   "Carrier_46_SpareInput(4_6)" AT %I2666.6 : Bool;   // SPARE INPUT
   "Carrier_46_SpareInput(4_7)" AT %I2666.7 : Bool;   // SPARE INPUT
   "Carrier_46_PB1_ProdHoldLH" AT %I2667.0 : Bool;   // PB 1 PRODUCTION HOLD LH
   "Carrier_46_PB2_ResetLH" AT %I2667.1 : Bool;   // PB 2 RESET LH
   "Carrier_46_PB3_ProdHoldRH" AT %I2667.2 : Bool;   // PB 3 PRODUCTION HOLD RH
   "Carrier_46_PB4_ResetRH" AT %I2667.3 : Bool;   // PB 4 RESET RH
   "Carrier_46_SpareInput(4_14)" AT %I2667.4 : Bool;   // SPARE INPUT
   "Carrier_46_SpareInput(4_15)" AT %I2667.5 : Bool;   // SPARE INPUT
   "Carrier_46_SpareInput(4_16)" AT %I2667.6 : Bool;   // SPARE INPUT
   "Carrier_46_SpareInput(4_17)" AT %I2667.7 : Bool;   // SPARE INPUT
   "Carrier_46_Slot5_Output" AT %IW2668 : Word;   // SLOT 5 OUTPUT WORD
   "Carrier_46_IRD400_HMI_24VDC_ENABLE" AT %I2668.0 : Bool;   // IRD 400 PANEL HMI 24V DC POWER
   "Carrier_46_FaultLight_LH" AT %I2668.1 : Bool;   // FAULT LIGHT LH
   "Carrier_46_RunLight_LH" AT %I2668.2 : Bool;   // RUN LIGHT LH
   "Carrier_46_FaultLight_RH" AT %I2668.3 : Bool;   // FAULT LIGHT RH
   "Carrier_46_RunLight_RH" AT %I2668.4 : Bool;   // RUN LIGHT RH
   "Carrier_46_SpareOutput(5_5)" AT %I2668.5 : Bool;   // SPARE OUTPUT
   "Carrier_46_SpareOutput(5_6)" AT %I2668.6 : Bool;   // SPARE OUTPUT
   "Carrier_46_SpareOutput(5_7)" AT %I2668.7 : Bool;   // SPARE OUTPUT
   "Carrier_46_ActualSpeed" AT %IW2670 : Word;   // ACTUAL SPEED
   "Carrier_46_CarrierDriveAlarm" AT %IW2672 : Word;   // CARRIER DRIVE ALARM
   "Carrier_46_CarrierDriveWarning" AT %IW2674 : Word;   // CARRIER DRIVE WARNING
   "Carrier_47_Status" AT %IW2700 : Word;   // CARRIER STATUS WORD
   "Carrier_47_Status.0" AT %I2700.0 : Bool;   // HEARTBEAT
   "Carrier_47_Status.1" AT %I2700.1 : Bool;   // MANUAL
   "Carrier_47_Status.2" AT %I2700.2 : Bool;   // IN_AUTO
   "Carrier_47_Status.3" AT %I2700.3 : Bool;   // POSITIONING_COMPLETE
   "Carrier_47_Status.4" AT %I2700.4 : Bool;   // PRODUCTION HOLD
   "Carrier_47_Status.5" AT %I2700.5 : Bool;   // CARRIER MOVING FORWARD
   "Carrier_47_Status.6" AT %I2700.6 : Bool;   // CARRIER MOVING REVERSE
   "Carrier_47_Status.7" AT %I2700.7 : Bool;   // CARRIER FAULT
   "Carrier_47_Status.8" AT %I2701.0 : Bool;   // CRASH DETECT TRIPPED
   "Carrier_47_Status.9" AT %I2701.1 : Bool;
   "Carrier_47_Status.10" AT %I2701.2 : Bool;
   "Carrier_47_Status.11" AT %I2701.3 : Bool;
   "Carrier_47_Status.12" AT %I2701.4 : Bool;
   "Carrier_47_Status.13" AT %I2701.5 : Bool;
   "Carrier_47_Status.14" AT %I2701.6 : Bool;
   "Carrier_47_Status.15" AT %I2701.7 : Bool;
   "Carrier_47_SDCFaultCode" AT %IW2702 : Word;   // SDC FAULT CODE
   "Carrier_47_CarrierPosition" AT %ID2704 : DWord;   // CARRIER POSITION
   "Carrier_47_CarrierNumber" AT %IW2708 : Word;   // CARRIER NUMBER
   "Carrier_47_G120DControlWord" AT %IW2710 : Word;   // G120D_STW1_CONTROL
   "Carrier_47_G120DControlWord.0" AT %I2710.0 : Bool;   // Bit_00_ON
   "Carrier_47_G120DControlWord.1" AT %I2710.1 : Bool;   // Bit_01_AUS2_INH
   "Carrier_47_G120DControlWord.2" AT %I2710.2 : Bool;   // Bit_02_AUS3_STOP
   "Carrier_47_G120DControlWord.3" AT %I2710.3 : Bool;   // Bit_03_EN
   "Carrier_47_G120DControlWord.4" AT %I2710.4 : Bool;   // Bit_04_EN_RAMP
   "Carrier_47_G120DControlWord.5" AT %I2710.5 : Bool;   // Bit_05_START_RAMP
   "Carrier_47_G120DControlWord.6" AT %I2710.6 : Bool;   // Bit_06_SETPOINT
   "Carrier_47_G120DControlWord.7" AT %I2710.7 : Bool;   // Bit_07_RESET
   "Carrier_47_G120DControlWord.8" AT %I2711.0 : Bool;   // Bit_08_JOG_R
   "Carrier_47_G120DControlWord.9" AT %I2711.1 : Bool;   // Bit_09_JOG_L
   "Carrier_47_G120DControlWord.10" AT %I2711.2 : Bool;   // Bit_10_CONTR_PLC
   "Carrier_47_G120DControlWord.11" AT %I2711.3 : Bool;   // Bit_11_REVERSE
   "Carrier_47_G120DControlWord.12" AT %I2711.4 : Bool;   // Bit_12_BRAKE_RELEASE
   "Carrier_47_G120DControlWord.13" AT %I2711.5 : Bool;   // Bit_13_DDS
   "Carrier_47_G120DControlWord.14" AT %I2711.6 : Bool;   // Bit_14_DO0
   "Carrier_47_G120DControlWord.15" AT %I2711.7 : Bool;   // Bit_15_DO1
   "Carrier_47_G120DStatusWord" AT %IW2712 : Word;   // G120D_ZSW1_STATUS
   "Carrier_47_G120DStatusWord.0" AT %I2712.0 : Bool;   // Bit_00_READY_RUN
   "Carrier_47_G120DStatusWord.1" AT %I2712.1 : Bool;   // Bit_01_READY_ON
   "Carrier_47_G120DStatusWord.2" AT %I2712.2 : Bool;   // Bit_02_ENABLE
   "Carrier_47_G120DStatusWord.3" AT %I2712.3 : Bool;   // Bit_03_FAULT
   "Carrier_47_G120DStatusWord.4" AT %I2712.4 : Bool;   // Bit_04_OFF2
   "Carrier_47_G120DStatusWord.5" AT %I2712.5 : Bool;   // Bit_05_OFF3
   "Carrier_47_G120DStatusWord.6" AT %I2712.6 : Bool;   // Bit_06_LOCK_OUT
   "Carrier_47_G120DStatusWord.7" AT %I2712.7 : Bool;   // Bit_07_WARN
   "Carrier_47_G120DStatusWord.8" AT %I2713.0 : Bool;   // Bit_08_NO_DEVIATION
   "Carrier_47_G120DStatusWord.9" AT %I2713.1 : Bool;   // Bit_09_CONTR_PLC
   "Carrier_47_G120DStatusWord.10" AT %I2713.2 : Bool;   // Bit_10_F_MAX
   "Carrier_47_G120DStatusWord.11" AT %I2713.3 : Bool;   // Bit_11_LIMIT_REACHED
   "Carrier_47_G120DStatusWord.12" AT %I2713.4 : Bool;   // Bit_12_BRAKE_OPEN
   "Carrier_47_G120DStatusWord.13" AT %I2713.5 : Bool;   // Bit_13_NO_OVERTEMP
   "Carrier_47_G120DStatusWord.14" AT %I2713.6 : Bool;   // Bit_14_CW_CCW
   "Carrier_47_G120DStatusWord.15" AT %I2713.7 : Bool;   // Bit_15_OVERL
   "Carrier_47_Slot2_Input" AT %IW2714 : Word;   // SLOT 2 INPUT WORD
   "Carrier_47_CrashDetectSW" AT %I2714.0 : Bool;   // CRASH DETECT SW
   "Carrier_47_SpareSafetyInput(2_1)" AT %I2714.1 : Bool;   // SPARE SAFETY INPUT
   "Carrier_47_SpareSafetyInput(2_2)" AT %I2714.2 : Bool;   // SPARE SAFETY INPUT
   "Carrier_47_SpareSafetyInput(2_3)" AT %I2714.3 : Bool;   // SPARE SAFETY INPUT
   "Carrier_47_SpareSafetyInput(2_4)" AT %I2714.4 : Bool;   // SPARE SAFETY INPUT
   "Carrier_47_SpareSafetyInput(2_5)" AT %I2714.5 : Bool;   // SPARE SAFETY INPUT
   "Carrier_47_SpareSafetyInput(2_6)" AT %I2714.6 : Bool;   // SPARE SAFETY INPUT
   "Carrier_47_SpareSafetyInput(2_7)" AT %I2714.7 : Bool;   // SPARE SAFETY INPUT
   "Carrier_47_Slot3_SafetyOutput" AT %IW2715 : Word;   // SLOT 3 SAFETY OUTPUT WORD
   "Carrier_47_Crash_Detect_OK" AT %I2715.0 : Bool;   // CARRIER CRASH DETECT
   "Carrier_47_SpareSafetyOutput(3_1)" AT %I2715.1 : Bool;   // SPARE SAFETY OUTPUT
   "Carrier_47_SpareSafetyOutput(3_2)" AT %I2715.2 : Bool;   // SPARE SAFETY OUTPUT
   "Carrier_47_SpareSafetyOutput(3_3)" AT %I2715.3 : Bool;   // SPARE SAFETY OUTPUT
   "Carrier_47_SpareSafetyOutput(3_4)" AT %I2715.4 : Bool;   // SPARE SAFETY OUTPUT
   "Carrier_47_SpareSafetyOutput(3_5)" AT %I2715.5 : Bool;   // SPARE SAFETY OUTPUT
   "Carrier_47_SpareSafetyOutput(3_6)" AT %I2715.6 : Bool;   // SPARE SAFETY OUTPUT
   "Carrier_47_SpareSafetyOutput(3_7)" AT %I2715.7 : Bool;   // SPARE SAFETY OUTPUT
   "Carrier_47_Slot4_Input" AT %IW2716 : Word;   // SLOT 4 INPUT WORD
   "Carrier_47_480VPowerOn_MDCB1" AT %I2716.0 : Bool;   // 480 VAC POWER ON MDCB 1
   "Carrier_47_SpareInput(4_1)" AT %I2716.1 : Bool;   // SPARE INPUT
   "Carrier_47_SpareInput(4_2)" AT %I2716.2 : Bool;   // SPARE INPUT
   "Carrier_47_SitopSelectStatus" AT %I2716.3 : Bool;   // SITOP SELECT STATUS
   "Carrier_47_DCsupplyOnPSCB2" AT %I2716.4 : Bool;   // DC SUPPLY ON PSCB 2
   "Carrier_47_SpareInput(4_5)" AT %I2716.5 : Bool;   // SPARE INPUT
   "Carrier_47_SpareInput(4_6)" AT %I2716.6 : Bool;   // SPARE INPUT
   "Carrier_47_SpareInput(4_7)" AT %I2716.7 : Bool;   // SPARE INPUT
   "Carrier_47_PB1_ProdHoldLH" AT %I2717.0 : Bool;   // PB 1 PRODUCTION HOLD LH
   "Carrier_47_PB2_ResetLH" AT %I2717.1 : Bool;   // PB 2 RESET LH
   "Carrier_47_PB3_ProdHoldRH" AT %I2717.2 : Bool;   // PB 3 PRODUCTION HOLD RH
   "Carrier_47_PB4_ResetRH" AT %I2717.3 : Bool;   // PB 4 RESET RH
   "Carrier_47_SpareInput(4_14)" AT %I2717.4 : Bool;   // SPARE INPUT
   "Carrier_47_SpareInput(4_15)" AT %I2717.5 : Bool;   // SPARE INPUT
   "Carrier_47_SpareInput(4_16)" AT %I2717.6 : Bool;   // SPARE INPUT
   "Carrier_47_SpareInput(4_17)" AT %I2717.7 : Bool;   // SPARE INPUT
   "Carrier_47_Slot5_Output" AT %IW2718 : Word;   // SLOT 5 OUTPUT WORD
   "Carrier_47_IRD400_HMI_24VDC_ENABLE" AT %I2718.0 : Bool;   // IRD 400 PANEL HMI 24V DC POWER
   "Carrier_47_FaultLight_LH" AT %I2718.1 : Bool;   // FAULT LIGHT LH
   "Carrier_47_RunLight_LH" AT %I2718.2 : Bool;   // RUN LIGHT LH
   "Carrier_47_FaultLight_RH" AT %I2718.3 : Bool;   // FAULT LIGHT RH
   "Carrier_47_RunLight_RH" AT %I2718.4 : Bool;   // RUN LIGHT RH
   "Carrier_47_SpareOutput(5_5)" AT %I2718.5 : Bool;   // SPARE OUTPUT
   "Carrier_47_SpareOutput(5_6)" AT %I2718.6 : Bool;   // SPARE OUTPUT
   "Carrier_47_SpareOutput(5_7)" AT %I2718.7 : Bool;   // SPARE OUTPUT
   "Carrier_47_ActualSpeed" AT %IW2720 : Word;   // ACTUAL SPEED
   "Carrier_47_CarrierDriveAlarm" AT %IW2722 : Word;   // CARRIER DRIVE ALARM
   "Carrier_47_CarrierDriveWarning" AT %IW2724 : Word;   // CARRIER DRIVE WARNING
   "Carrier_48_Status" AT %IW2750 : Word;   // CARRIER STATUS WORD
   "Carrier_48_Status.0" AT %I2750.0 : Bool;   // HEARTBEAT
   "Carrier_48_Status.1" AT %I2750.1 : Bool;   // MANUAL
   "Carrier_48_Status.2" AT %I2750.2 : Bool;   // IN_AUTO
   "Carrier_48_Status.3" AT %I2750.3 : Bool;   // POSITIONING_COMPLETE
   "Carrier_48_Status.4" AT %I2750.4 : Bool;   // PRODUCTION HOLD
   "Carrier_48_Status.5" AT %I2750.5 : Bool;   // CARRIER MOVING FORWARD
   "Carrier_48_Status.6" AT %I2750.6 : Bool;   // CARRIER MOVING REVERSE
   "Carrier_48_Status.7" AT %I2750.7 : Bool;   // CARRIER FAULT
   "Carrier_48_Status.8" AT %I2751.0 : Bool;   // CRASH DETECT TRIPPED
   "Carrier_48_Status.9" AT %I2751.1 : Bool;
   "Carrier_48_Status.10" AT %I2751.2 : Bool;
   "Carrier_48_Status.11" AT %I2751.3 : Bool;
   "Carrier_48_Status.12" AT %I2751.4 : Bool;
   "Carrier_48_Status.13" AT %I2751.5 : Bool;
   "Carrier_48_Status.14" AT %I2751.6 : Bool;
   "Carrier_48_Status.15" AT %I2751.7 : Bool;
   "Carrier_48_SDCFaultCode" AT %IW2752 : Word;   // SDC FAULT CODE
   "Carrier_48_CarrierPosition" AT %ID2754 : DWord;   // CARRIER POSITION
   "Carrier_48_CarrierNumber" AT %IW2758 : Word;   // CARRIER NUMBER
   "Carrier_48_G120DControlWord" AT %IW2760 : Word;   // G120D_STW1_CONTROL
   "Carrier_48_G120DControlWord.0" AT %I2760.0 : Bool;   // Bit_00_ON
   "Carrier_48_G120DControlWord.1" AT %I2760.1 : Bool;   // Bit_01_AUS2_INH
   "Carrier_48_G120DControlWord.2" AT %I2760.2 : Bool;   // Bit_02_AUS3_STOP
   "Carrier_48_G120DControlWord.3" AT %I2760.3 : Bool;   // Bit_03_EN
   "Carrier_48_G120DControlWord.4" AT %I2760.4 : Bool;   // Bit_04_EN_RAMP
   "Carrier_48_G120DControlWord.5" AT %I2760.5 : Bool;   // Bit_05_START_RAMP
   "Carrier_48_G120DControlWord.6" AT %I2760.6 : Bool;   // Bit_06_SETPOINT
   "Carrier_48_G120DControlWord.7" AT %I2760.7 : Bool;   // Bit_07_RESET
   "Carrier_48_G120DControlWord.8" AT %I2761.0 : Bool;   // Bit_08_JOG_R
   "Carrier_48_G120DControlWord.9" AT %I2761.1 : Bool;   // Bit_09_JOG_L
   "Carrier_48_G120DControlWord.10" AT %I2761.2 : Bool;   // Bit_10_CONTR_PLC
   "Carrier_48_G120DControlWord.11" AT %I2761.3 : Bool;   // Bit_11_REVERSE
   "Carrier_48_G120DControlWord.12" AT %I2761.4 : Bool;   // Bit_12_BRAKE_RELEASE
   "Carrier_48_G120DControlWord.13" AT %I2761.5 : Bool;   // Bit_13_DDS
   "Carrier_48_G120DControlWord.14" AT %I2761.6 : Bool;   // Bit_14_DO0
   "Carrier_48_G120DControlWord.15" AT %I2761.7 : Bool;   // Bit_15_DO1
   "Carrier_48_G120DStatusWord" AT %IW2762 : Word;   // G120D_ZSW1_STATUS
   "Carrier_48_G120DStatusWord.0" AT %I2762.0 : Bool;   // Bit_00_READY_RUN
   "Carrier_48_G120DStatusWord.1" AT %I2762.1 : Bool;   // Bit_01_READY_ON
   "Carrier_48_G120DStatusWord.2" AT %I2762.2 : Bool;   // Bit_02_ENABLE
   "Carrier_48_G120DStatusWord.3" AT %I2762.3 : Bool;   // Bit_03_FAULT
   "Carrier_48_G120DStatusWord.4" AT %I2762.4 : Bool;   // Bit_04_OFF2
   "Carrier_48_G120DStatusWord.5" AT %I2762.5 : Bool;   // Bit_05_OFF3
   "Carrier_48_G120DStatusWord.6" AT %I2762.6 : Bool;   // Bit_06_LOCK_OUT
   "Carrier_48_G120DStatusWord.7" AT %I2762.7 : Bool;   // Bit_07_WARN
   "Carrier_48_G120DStatusWord.8" AT %I2763.0 : Bool;   // Bit_08_NO_DEVIATION
   "Carrier_48_G120DStatusWord.9" AT %I2763.1 : Bool;   // Bit_09_CONTR_PLC
   "Carrier_48_G120DStatusWord.10" AT %I2763.2 : Bool;   // Bit_10_F_MAX
   "Carrier_48_G120DStatusWord.11" AT %I2763.3 : Bool;   // Bit_11_LIMIT_REACHED
   "Carrier_48_G120DStatusWord.12" AT %I2763.4 : Bool;   // Bit_12_BRAKE_OPEN
   "Carrier_48_G120DStatusWord.13" AT %I2763.5 : Bool;   // Bit_13_NO_OVERTEMP
   "Carrier_48_G120DStatusWord.14" AT %I2763.6 : Bool;   // Bit_14_CW_CCW
   "Carrier_48_G120DStatusWord.15" AT %I2763.7 : Bool;   // Bit_15_OVERL
   "Carrier_48_Slot2_Input" AT %IW2764 : Word;   // SLOT 2 INPUT WORD
   "Carrier_48_CrashDetectSW" AT %I2764.0 : Bool;   // CRASH DETECT SW
   "Carrier_48_SpareSafetyInput(2_1)" AT %I2764.1 : Bool;   // SPARE SAFETY INPUT
   "Carrier_48_SpareSafetyInput(2_2)" AT %I2764.2 : Bool;   // SPARE SAFETY INPUT
   "Carrier_48_SpareSafetyInput(2_3)" AT %I2764.3 : Bool;   // SPARE SAFETY INPUT
   "Carrier_48_SpareSafetyInput(2_4)" AT %I2764.4 : Bool;   // SPARE SAFETY INPUT
   "Carrier_48_SpareSafetyInput(2_5)" AT %I2764.5 : Bool;   // SPARE SAFETY INPUT
   "Carrier_48_SpareSafetyInput(2_6)" AT %I2764.6 : Bool;   // SPARE SAFETY INPUT
   "Carrier_48_SpareSafetyInput(2_7)" AT %I2764.7 : Bool;   // SPARE SAFETY INPUT
   "Carrier_48_Slot3_SafetyOutput" AT %IW2765 : Word;   // SLOT 3 SAFETY OUTPUT WORD
   "Carrier_48_Crash_Detect_OK" AT %I2765.0 : Bool;   // CARRIER CRASH DETECT
   "Carrier_48_SpareSafetyOutput(3_1)" AT %I2765.1 : Bool;   // SPARE SAFETY OUTPUT
   "Carrier_48_SpareSafetyOutput(3_2)" AT %I2765.2 : Bool;   // SPARE SAFETY OUTPUT
   "Carrier_48_SpareSafetyOutput(3_3)" AT %I2765.3 : Bool;   // SPARE SAFETY OUTPUT
   "Carrier_48_SpareSafetyOutput(3_4)" AT %I2765.4 : Bool;   // SPARE SAFETY OUTPUT
   "Carrier_48_SpareSafetyOutput(3_5)" AT %I2765.5 : Bool;   // SPARE SAFETY OUTPUT
   "Carrier_48_SpareSafetyOutput(3_6)" AT %I2765.6 : Bool;   // SPARE SAFETY OUTPUT
   "Carrier_48_SpareSafetyOutput(3_7)" AT %I2765.7 : Bool;   // SPARE SAFETY OUTPUT
   "Carrier_48_Slot4_Input" AT %IW2766 : Word;   // SLOT 4 INPUT WORD
   "Carrier_48_480VPowerOn_MDCB1" AT %I2766.0 : Bool;   // 480 VAC POWER ON MDCB 1
   "Carrier_48_SpareInput(4_1)" AT %I2766.1 : Bool;   // SPARE INPUT
   "Carrier_48_SpareInput(4_2)" AT %I2766.2 : Bool;   // SPARE INPUT
   "Carrier_48_SitopSelectStatus" AT %I2766.3 : Bool;   // SITOP SELECT STATUS
   "Carrier_48_DCsupplyOnPSCB2" AT %I2766.4 : Bool;   // DC SUPPLY ON PSCB 2
   "Carrier_48_SpareInput(4_5)" AT %I2766.5 : Bool;   // SPARE INPUT
   "Carrier_48_SpareInput(4_6)" AT %I2766.6 : Bool;   // SPARE INPUT
   "Carrier_48_SpareInput(4_7)" AT %I2766.7 : Bool;   // SPARE INPUT
   "Carrier_48_PB1_ProdHoldLH" AT %I2767.0 : Bool;   // PB 1 PRODUCTION HOLD LH
   "Carrier_48_PB2_ResetLH" AT %I2767.1 : Bool;   // PB 2 RESET LH
   "Carrier_48_PB3_ProdHoldRH" AT %I2767.2 : Bool;   // PB 3 PRODUCTION HOLD RH
   "Carrier_48_PB4_ResetRH" AT %I2767.3 : Bool;   // PB 4 RESET RH
   "Carrier_48_SpareInput(4_14)" AT %I2767.4 : Bool;   // SPARE INPUT
   "Carrier_48_SpareInput(4_15)" AT %I2767.5 : Bool;   // SPARE INPUT
   "Carrier_48_SpareInput(4_16)" AT %I2767.6 : Bool;   // SPARE INPUT
   "Carrier_48_SpareInput(4_17)" AT %I2767.7 : Bool;   // SPARE INPUT
   "Carrier_48_Slot5_Output" AT %IW2768 : Word;   // SLOT 5 OUTPUT WORD
   "Carrier_48_IRD400_HMI_24VDC_ENABLE" AT %I2768.0 : Bool;   // IRD 400 PANEL HMI 24V DC POWER
   "Carrier_48_FaultLight_LH" AT %I2768.1 : Bool;   // FAULT LIGHT LH
   "Carrier_48_RunLight_LH" AT %I2768.2 : Bool;   // RUN LIGHT LH
   "Carrier_48_FaultLight_RH" AT %I2768.3 : Bool;   // FAULT LIGHT RH
   "Carrier_48_RunLight_RH" AT %I2768.4 : Bool;   // RUN LIGHT RH
   "Carrier_48_SpareOutput(5_5)" AT %I2768.5 : Bool;   // SPARE OUTPUT
   "Carrier_48_SpareOutput(5_6)" AT %I2768.6 : Bool;   // SPARE OUTPUT
   "Carrier_48_SpareOutput(5_7)" AT %I2768.7 : Bool;   // SPARE OUTPUT
   "Carrier_48_ActualSpeed" AT %IW2770 : Word;   // ACTUAL SPEED
   "Carrier_48_CarrierDriveAlarm" AT %IW2772 : Word;   // CARRIER DRIVE ALARM
   "Carrier_48_CarrierDriveWarning" AT %IW2774 : Word;   // CARRIER DRIVE WARNING
   "Carrier_49_Status" AT %IW2800 : Word;   // CARRIER STATUS WORD
   "Carrier_49_Status.0" AT %I2800.0 : Bool;   // HEARTBEAT
   "Carrier_49_Status.1" AT %I2800.1 : Bool;   // MANUAL
   "Carrier_49_Status.2" AT %I2800.2 : Bool;   // IN_AUTO
   "Carrier_49_Status.3" AT %I2800.3 : Bool;   // POSITIONING_COMPLETE
   "Carrier_49_Status.4" AT %I2800.4 : Bool;   // PRODUCTION HOLD
   "Carrier_49_Status.5" AT %I2800.5 : Bool;   // CARRIER MOVING FORWARD
   "Carrier_49_Status.6" AT %I2800.6 : Bool;   // CARRIER MOVING REVERSE
   "Carrier_49_Status.7" AT %I2800.7 : Bool;   // CARRIER FAULT
   "Carrier_49_Status.8" AT %I2801.0 : Bool;   // CRASH DETECT TRIPPED
   "Carrier_49_Status.9" AT %I2801.1 : Bool;
   "Carrier_49_Status.10" AT %I2801.2 : Bool;
   "Carrier_49_Status.11" AT %I2801.3 : Bool;
   "Carrier_49_Status.12" AT %I2801.4 : Bool;
   "Carrier_49_Status.13" AT %I2801.5 : Bool;
   "Carrier_49_Status.14" AT %I2801.6 : Bool;
   "Carrier_49_Status.15" AT %I2801.7 : Bool;
   "Carrier_49_SDCFaultCode" AT %IW2802 : Word;   // SDC FAULT CODE
   "Carrier_49_CarrierPosition" AT %ID2804 : DWord;   // CARRIER POSITION
   "Carrier_49_CarrierNumber" AT %IW2808 : Word;   // CARRIER NUMBER
   "Carrier_49_G120DControlWord" AT %IW2810 : Word;   // G120D_STW1_CONTROL
   "Carrier_49_G120DControlWord.0" AT %I2810.0 : Bool;   // Bit_00_ON
   "Carrier_49_G120DControlWord.1" AT %I2810.1 : Bool;   // Bit_01_AUS2_INH
   "Carrier_49_G120DControlWord.2" AT %I2810.2 : Bool;   // Bit_02_AUS3_STOP
   "Carrier_49_G120DControlWord.3" AT %I2810.3 : Bool;   // Bit_03_EN
   "Carrier_49_G120DControlWord.4" AT %I2810.4 : Bool;   // Bit_04_EN_RAMP
   "Carrier_49_G120DControlWord.5" AT %I2810.5 : Bool;   // Bit_05_START_RAMP
   "Carrier_49_G120DControlWord.6" AT %I2810.6 : Bool;   // Bit_06_SETPOINT
   "Carrier_49_G120DControlWord.7" AT %I2810.7 : Bool;   // Bit_07_RESET
   "Carrier_49_G120DControlWord.8" AT %I2811.0 : Bool;   // Bit_08_JOG_R
   "Carrier_49_G120DControlWord.9" AT %I2811.1 : Bool;   // Bit_09_JOG_L
   "Carrier_49_G120DControlWord.10" AT %I2811.2 : Bool;   // Bit_10_CONTR_PLC
   "Carrier_49_G120DControlWord.11" AT %I2811.3 : Bool;   // Bit_11_REVERSE
   "Carrier_49_G120DControlWord.12" AT %I2811.4 : Bool;   // Bit_12_BRAKE_RELEASE
   "Carrier_49_G120DControlWord.13" AT %I2811.5 : Bool;   // Bit_13_DDS
   "Carrier_49_G120DControlWord.14" AT %I2811.6 : Bool;   // Bit_14_DO0
   "Carrier_49_G120DControlWord.15" AT %I2811.7 : Bool;   // Bit_15_DO1
   "Carrier_49_G120DStatusWord" AT %IW2812 : Word;   // G120D_ZSW1_STATUS
   "Carrier_49_G120DStatusWord.0" AT %I2812.0 : Bool;   // Bit_00_READY_RUN
   "Carrier_49_G120DStatusWord.1" AT %I2812.1 : Bool;   // Bit_01_READY_ON
   "Carrier_49_G120DStatusWord.2" AT %I2812.2 : Bool;   // Bit_02_ENABLE
   "Carrier_49_G120DStatusWord.3" AT %I2812.3 : Bool;   // Bit_03_FAULT
   "Carrier_49_G120DStatusWord.4" AT %I2812.4 : Bool;   // Bit_04_OFF2
   "Carrier_49_G120DStatusWord.5" AT %I2812.5 : Bool;   // Bit_05_OFF3
   "Carrier_49_G120DStatusWord.6" AT %I2812.6 : Bool;   // Bit_06_LOCK_OUT
   "Carrier_49_G120DStatusWord.7" AT %I2812.7 : Bool;   // Bit_07_WARN
   "Carrier_49_G120DStatusWord.8" AT %I2813.0 : Bool;   // Bit_08_NO_DEVIATION
   "Carrier_49_G120DStatusWord.9" AT %I2813.1 : Bool;   // Bit_09_CONTR_PLC
   "Carrier_49_G120DStatusWord.10" AT %I2813.2 : Bool;   // Bit_10_F_MAX
   "Carrier_49_G120DStatusWord.11" AT %I2813.3 : Bool;   // Bit_11_LIMIT_REACHED
   "Carrier_49_G120DStatusWord.12" AT %I2813.4 : Bool;   // Bit_12_BRAKE_OPEN
   "Carrier_49_G120DStatusWord.13" AT %I2813.5 : Bool;   // Bit_13_NO_OVERTEMP
   "Carrier_49_G120DStatusWord.14" AT %I2813.6 : Bool;   // Bit_14_CW_CCW
   "Carrier_49_G120DStatusWord.15" AT %I2813.7 : Bool;   // Bit_15_OVERL
   "Carrier_49_Slot2_Input" AT %IW2814 : Word;   // SLOT 2 INPUT WORD
   "Carrier_49_CrashDetectSW" AT %I2814.0 : Bool;   // CRASH DETECT SW
   "Carrier_49_SpareSafetyInput(2_1)" AT %I2814.1 : Bool;   // SPARE SAFETY INPUT
   "Carrier_49_SpareSafetyInput(2_2)" AT %I2814.2 : Bool;   // SPARE SAFETY INPUT
   "Carrier_49_SpareSafetyInput(2_3)" AT %I2814.3 : Bool;   // SPARE SAFETY INPUT
   "Carrier_49_SpareSafetyInput(2_4)" AT %I2814.4 : Bool;   // SPARE SAFETY INPUT
   "Carrier_49_SpareSafetyInput(2_5)" AT %I2814.5 : Bool;   // SPARE SAFETY INPUT
   "Carrier_49_SpareSafetyInput(2_6)" AT %I2814.6 : Bool;   // SPARE SAFETY INPUT
   "Carrier_49_SpareSafetyInput(2_7)" AT %I2814.7 : Bool;   // SPARE SAFETY INPUT
   "Carrier_49_Slot3_SafetyOutput" AT %IW2815 : Word;   // SLOT 3 SAFETY OUTPUT WORD
   "Carrier_49_Crash_Detect_OK" AT %I2815.0 : Bool;   // CARRIER CRASH DETECT
   "Carrier_49_SpareSafetyOutput(3_1)" AT %I2815.1 : Bool;   // SPARE SAFETY OUTPUT
   "Carrier_49_SpareSafetyOutput(3_2)" AT %I2815.2 : Bool;   // SPARE SAFETY OUTPUT
   "Carrier_49_SpareSafetyOutput(3_3)" AT %I2815.3 : Bool;   // SPARE SAFETY OUTPUT
   "Carrier_49_SpareSafetyOutput(3_4)" AT %I2815.4 : Bool;   // SPARE SAFETY OUTPUT
   "Carrier_49_SpareSafetyOutput(3_5)" AT %I2815.5 : Bool;   // SPARE SAFETY OUTPUT
   "Carrier_49_SpareSafetyOutput(3_6)" AT %I2815.6 : Bool;   // SPARE SAFETY OUTPUT
   "Carrier_49_SpareSafetyOutput(3_7)" AT %I2815.7 : Bool;   // SPARE SAFETY OUTPUT
   "Carrier_49_Slot4_Input" AT %IW2816 : Word;   // SLOT 4 INPUT WORD
   "Carrier_49_480VPowerOn_MDCB1" AT %I2816.0 : Bool;   // 480 VAC POWER ON MDCB 1
   "Carrier_49_SpareInput(4_1)" AT %I2816.1 : Bool;   // SPARE INPUT
   "Carrier_49_SpareInput(4_2)" AT %I2816.2 : Bool;   // SPARE INPUT
   "Carrier_49_SitopSelectStatus" AT %I2816.3 : Bool;   // SITOP SELECT STATUS
   "Carrier_49_DCsupplyOnPSCB2" AT %I2816.4 : Bool;   // DC SUPPLY ON PSCB 2
   "Carrier_49_SpareInput(4_5)" AT %I2816.5 : Bool;   // SPARE INPUT
   "Carrier_49_SpareInput(4_6)" AT %I2816.6 : Bool;   // SPARE INPUT
   "Carrier_49_SpareInput(4_7)" AT %I2816.7 : Bool;   // SPARE INPUT
   "Carrier_49_PB1_ProdHoldLH" AT %I2817.0 : Bool;   // PB 1 PRODUCTION HOLD LH
   "Carrier_49_PB2_ResetLH" AT %I2817.1 : Bool;   // PB 2 RESET LH
   "Carrier_49_PB3_ProdHoldRH" AT %I2817.2 : Bool;   // PB 3 PRODUCTION HOLD RH
   "Carrier_49_PB4_ResetRH" AT %I2817.3 : Bool;   // PB 4 RESET RH
   "Carrier_49_SpareInput(4_14)" AT %I2817.4 : Bool;   // SPARE INPUT
   "Carrier_49_SpareInput(4_15)" AT %I2817.5 : Bool;   // SPARE INPUT
   "Carrier_49_SpareInput(4_16)" AT %I2817.6 : Bool;   // SPARE INPUT
   "Carrier_49_SpareInput(4_17)" AT %I2817.7 : Bool;   // SPARE INPUT
   "Carrier_49_Slot5_Output" AT %IW2818 : Word;   // SLOT 5 OUTPUT WORD
   "Carrier_49_IRD400_HMI_24VDC_ENABLE" AT %I2818.0 : Bool;   // IRD 400 PANEL HMI 24V DC POWER
   "Carrier_49_FaultLight_LH" AT %I2818.1 : Bool;   // FAULT LIGHT LH
   "Carrier_49_RunLight_LH" AT %I2818.2 : Bool;   // RUN LIGHT LH
   "Carrier_49_FaultLight_RH" AT %I2818.3 : Bool;   // FAULT LIGHT RH
   "Carrier_49_RunLight_RH" AT %I2818.4 : Bool;   // RUN LIGHT RH
   "Carrier_49_SpareOutput(5_5)" AT %I2818.5 : Bool;   // SPARE OUTPUT
   "Carrier_49_SpareOutput(5_6)" AT %I2818.6 : Bool;   // SPARE OUTPUT
   "Carrier_49_SpareOutput(5_7)" AT %I2818.7 : Bool;   // SPARE OUTPUT
   "Carrier_49_ActualSpeed" AT %IW2820 : Word;   // ACTUAL SPEED
   "Carrier_49_CarrierDriveAlarm" AT %IW2822 : Word;   // CARRIER DRIVE ALARM
   "Carrier_49_CarrierDriveWarning" AT %IW2824 : Word;   // CARRIER DRIVE WARNING
   "Carrier_50_Status" AT %IW2850 : Word;   // CARRIER STATUS WORD
   "Carrier_50_Status.0" AT %I2850.0 : Bool;   // HEARTBEAT
   "Carrier_50_Status.1" AT %I2850.1 : Bool;   // MANUAL
   "Carrier_50_Status.2" AT %I2850.2 : Bool;   // IN_AUTO
   "Carrier_50_Status.3" AT %I2850.3 : Bool;   // POSITIONING_COMPLETE
   "Carrier_50_Status.4" AT %I2850.4 : Bool;   // PRODUCTION HOLD
   "Carrier_50_Status.5" AT %I2850.5 : Bool;   // CARRIER MOVING FORWARD
   "Carrier_50_Status.6" AT %I2850.6 : Bool;   // CARRIER MOVING REVERSE
   "Carrier_50_Status.7" AT %I2850.7 : Bool;   // CARRIER FAULT
   "Carrier_50_Status.8" AT %I2851.0 : Bool;   // CRASH DETECT TRIPPED
   "Carrier_50_Status.9" AT %I2851.1 : Bool;
   "Carrier_50_Status.10" AT %I2851.2 : Bool;
   "Carrier_50_Status.11" AT %I2851.3 : Bool;
   "Carrier_50_Status.12" AT %I2851.4 : Bool;
   "Carrier_50_Status.13" AT %I2851.5 : Bool;
   "Carrier_50_Status.14" AT %I2851.6 : Bool;
   "Carrier_50_Status.15" AT %I2851.7 : Bool;
   "Carrier_50_SDCFaultCode" AT %IW2852 : Word;   // SDC FAULT CODE
   "Carrier_50_CarrierPosition" AT %ID2854 : DWord;   // CARRIER POSITION
   "Carrier_50_CarrierNumber" AT %IW2858 : Word;   // CARRIER NUMBER
   "Carrier_50_G120DControlWord" AT %IW2860 : Word;   // G120D_STW1_CONTROL
   "Carrier_50_G120DControlWord.0" AT %I2860.0 : Bool;   // Bit_00_ON
   "Carrier_50_G120DControlWord.1" AT %I2860.1 : Bool;   // Bit_01_AUS2_INH
   "Carrier_50_G120DControlWord.2" AT %I2860.2 : Bool;   // Bit_02_AUS3_STOP
   "Carrier_50_G120DControlWord.3" AT %I2860.3 : Bool;   // Bit_03_EN
   "Carrier_50_G120DControlWord.4" AT %I2860.4 : Bool;   // Bit_04_EN_RAMP
   "Carrier_50_G120DControlWord.5" AT %I2860.5 : Bool;   // Bit_05_START_RAMP
   "Carrier_50_G120DControlWord.6" AT %I2860.6 : Bool;   // Bit_06_SETPOINT
   "Carrier_50_G120DControlWord.7" AT %I2860.7 : Bool;   // Bit_07_RESET
   "Carrier_50_G120DControlWord.8" AT %I2861.0 : Bool;   // Bit_08_JOG_R
   "Carrier_50_G120DControlWord.9" AT %I2861.1 : Bool;   // Bit_09_JOG_L
   "Carrier_50_G120DControlWord.10" AT %I2861.2 : Bool;   // Bit_10_CONTR_PLC
   "Carrier_50_G120DControlWord.11" AT %I2861.3 : Bool;   // Bit_11_REVERSE
   "Carrier_50_G120DControlWord.12" AT %I2861.4 : Bool;   // Bit_12_BRAKE_RELEASE
   "Carrier_50_G120DControlWord.13" AT %I2861.5 : Bool;   // Bit_13_DDS
   "Carrier_50_G120DControlWord.14" AT %I2861.6 : Bool;   // Bit_14_DO0
   "Carrier_50_G120DControlWord.15" AT %I2861.7 : Bool;   // Bit_15_DO1
   "Carrier_50_G120DStatusWord" AT %IW2862 : Word;   // G120D_ZSW1_STATUS
   "Carrier_50_G120DStatusWord.0" AT %I2862.0 : Bool;   // Bit_00_READY_RUN
   "Carrier_50_G120DStatusWord.1" AT %I2862.1 : Bool;   // Bit_01_READY_ON
   "Carrier_50_G120DStatusWord.2" AT %I2862.2 : Bool;   // Bit_02_ENABLE
   "Carrier_50_G120DStatusWord.3" AT %I2862.3 : Bool;   // Bit_03_FAULT
   "Carrier_50_G120DStatusWord.4" AT %I2862.4 : Bool;   // Bit_04_OFF2
   "Carrier_50_G120DStatusWord.5" AT %I2862.5 : Bool;   // Bit_05_OFF3
   "Carrier_50_G120DStatusWord.6" AT %I2862.6 : Bool;   // Bit_06_LOCK_OUT
   "Carrier_50_G120DStatusWord.7" AT %I2862.7 : Bool;   // Bit_07_WARN
   "Carrier_50_G120DStatusWord.8" AT %I2863.0 : Bool;   // Bit_08_NO_DEVIATION
   "Carrier_50_G120DStatusWord.9" AT %I2863.1 : Bool;   // Bit_09_CONTR_PLC
   "Carrier_50_G120DStatusWord.10" AT %I2863.2 : Bool;   // Bit_10_F_MAX
   "Carrier_50_G120DStatusWord.11" AT %I2863.3 : Bool;   // Bit_11_LIMIT_REACHED
   "Carrier_50_G120DStatusWord.12" AT %I2863.4 : Bool;   // Bit_12_BRAKE_OPEN
   "Carrier_50_G120DStatusWord.13" AT %I2863.5 : Bool;   // Bit_13_NO_OVERTEMP
   "Carrier_50_G120DStatusWord.14" AT %I2863.6 : Bool;   // Bit_14_CW_CCW
   "Carrier_50_G120DStatusWord.15" AT %I2863.7 : Bool;   // Bit_15_OVERL
   "Carrier_50_Slot2_Input" AT %IW2864 : Word;   // SLOT 2 INPUT WORD
   "Carrier_50_CrashDetectSW" AT %I2864.0 : Bool;   // CRASH DETECT SW
   "Carrier_50_SpareSafetyInput(2_1)" AT %I2864.1 : Bool;   // SPARE SAFETY INPUT
   "Carrier_50_SpareSafetyInput(2_2)" AT %I2864.2 : Bool;   // SPARE SAFETY INPUT
   "Carrier_50_SpareSafetyInput(2_3)" AT %I2864.3 : Bool;   // SPARE SAFETY INPUT
   "Carrier_50_SpareSafetyInput(2_4)" AT %I2864.4 : Bool;   // SPARE SAFETY INPUT
   "Carrier_50_SpareSafetyInput(2_5)" AT %I2864.5 : Bool;   // SPARE SAFETY INPUT
   "Carrier_50_SpareSafetyInput(2_6)" AT %I2864.6 : Bool;   // SPARE SAFETY INPUT
   "Carrier_50_SpareSafetyInput(2_7)" AT %I2864.7 : Bool;   // SPARE SAFETY INPUT
   "Carrier_50_Slot3_SafetyOutput" AT %IW2865 : Word;   // SLOT 3 SAFETY OUTPUT WORD
   "Carrier_50_Crash_Detect_OK" AT %I2865.0 : Bool;   // CARRIER CRASH DETECT
   "Carrier_50_SpareSafetyOutput(3_1)" AT %I2865.1 : Bool;   // SPARE SAFETY OUTPUT
   "Carrier_50_SpareSafetyOutput(3_2)" AT %I2865.2 : Bool;   // SPARE SAFETY OUTPUT
   "Carrier_50_SpareSafetyOutput(3_3)" AT %I2865.3 : Bool;   // SPARE SAFETY OUTPUT
   "Carrier_50_SpareSafetyOutput(3_4)" AT %I2865.4 : Bool;   // SPARE SAFETY OUTPUT
   "Carrier_50_SpareSafetyOutput(3_5)" AT %I2865.5 : Bool;   // SPARE SAFETY OUTPUT
   "Carrier_50_SpareSafetyOutput(3_6)" AT %I2865.6 : Bool;   // SPARE SAFETY OUTPUT
   "Carrier_50_SpareSafetyOutput(3_7)" AT %I2865.7 : Bool;   // SPARE SAFETY OUTPUT
   "Carrier_50_Slot4_Input" AT %IW2866 : Word;   // SLOT 4 INPUT WORD
   "Carrier_50_480VPowerOn_MDCB1" AT %I2866.0 : Bool;   // 480 VAC POWER ON MDCB 1
   "Carrier_50_SpareInput(4_1)" AT %I2866.1 : Bool;   // SPARE INPUT
   "Carrier_50_SpareInput(4_2)" AT %I2866.2 : Bool;   // SPARE INPUT
   "Carrier_50_SitopSelectStatus" AT %I2866.3 : Bool;   // SITOP SELECT STATUS
   "Carrier_50_DCsupplyOnPSCB2" AT %I2866.4 : Bool;   // DC SUPPLY ON PSCB 2
   "Carrier_50_SpareInput(4_5)" AT %I2866.5 : Bool;   // SPARE INPUT
   "Carrier_50_SpareInput(4_6)" AT %I2866.6 : Bool;   // SPARE INPUT
   "Carrier_50_SpareInput(4_7)" AT %I2866.7 : Bool;   // SPARE INPUT
   "Carrier_50_PB1_ProdHoldLH" AT %I2867.0 : Bool;   // PB 1 PRODUCTION HOLD LH
   "Carrier_50_PB2_ResetLH" AT %I2867.1 : Bool;   // PB 2 RESET LH
   "Carrier_50_PB3_ProdHoldRH" AT %I2867.2 : Bool;   // PB 3 PRODUCTION HOLD RH
   "Carrier_50_PB4_ResetRH" AT %I2867.3 : Bool;   // PB 4 RESET RH
   "Carrier_50_SpareInput(4_14)" AT %I2867.4 : Bool;   // SPARE INPUT
   "Carrier_50_SpareInput(4_15)" AT %I2867.5 : Bool;   // SPARE INPUT
   "Carrier_50_SpareInput(4_16)" AT %I2867.6 : Bool;   // SPARE INPUT
   "Carrier_50_SpareInput(4_17)" AT %I2867.7 : Bool;   // SPARE INPUT
   "Carrier_50_Slot5_Output" AT %IW2868 : Word;   // SLOT 5 OUTPUT WORD
   "Carrier_50_IRD400_HMI_24VDC_ENABLE" AT %I2868.0 : Bool;   // IRD 400 PANEL HMI 24V DC POWER
   "Carrier_50_FaultLight_LH" AT %I2868.1 : Bool;   // FAULT LIGHT LH
   "Carrier_50_RunLight_LH" AT %I2868.2 : Bool;   // RUN LIGHT LH
   "Carrier_50_FaultLight_RH" AT %I2868.3 : Bool;   // FAULT LIGHT RH
   "Carrier_50_RunLight_RH" AT %I2868.4 : Bool;   // RUN LIGHT RH
   "Carrier_50_SpareOutput(5_5)" AT %I2868.5 : Bool;   // SPARE OUTPUT
   "Carrier_50_SpareOutput(5_6)" AT %I2868.6 : Bool;   // SPARE OUTPUT
   "Carrier_50_SpareOutput(5_7)" AT %I2868.7 : Bool;   // SPARE OUTPUT
   "Carrier_50_ActualSpeed" AT %IW2870 : Word;   // ACTUAL SPEED
   "Carrier_50_CarrierDriveAlarm" AT %IW2872 : Word;   // CARRIER DRIVE ALARM
   "Carrier_50_CarrierDriveWarning" AT %IW2874 : Word;   // CARRIER DRIVE WARNING
   "Carrier_51_Status" AT %IW2900 : Word;   // CARRIER STATUS WORD
   "Carrier_51_Status.0" AT %I2900.0 : Bool;   // HEARTBEAT
   "Carrier_51_Status.1" AT %I2900.1 : Bool;   // MANUAL
   "Carrier_51_Status.2" AT %I2900.2 : Bool;   // IN_AUTO
   "Carrier_51_Status.3" AT %I2900.3 : Bool;   // POSITIONING_COMPLETE
   "Carrier_51_Status.4" AT %I2900.4 : Bool;   // PRODUCTION HOLD
   "Carrier_51_Status.5" AT %I2900.5 : Bool;   // CARRIER MOVING FORWARD
   "Carrier_51_Status.6" AT %I2900.6 : Bool;   // CARRIER MOVING REVERSE
   "Carrier_51_Status.7" AT %I2900.7 : Bool;   // CARRIER FAULT
   "Carrier_51_Status.8" AT %I2901.0 : Bool;   // CRASH DETECT TRIPPED
   "Carrier_51_Status.9" AT %I2901.1 : Bool;
   "Carrier_51_Status.10" AT %I2901.2 : Bool;
   "Carrier_51_Status.11" AT %I2901.3 : Bool;
   "Carrier_51_Status.12" AT %I2901.4 : Bool;
   "Carrier_51_Status.13" AT %I2901.5 : Bool;
   "Carrier_51_Status.14" AT %I2901.6 : Bool;
   "Carrier_51_Status.15" AT %I2901.7 : Bool;
   "Carrier_51_SDCFaultCode" AT %IW2902 : Word;   // SDC FAULT CODE
   "Carrier_51_CarrierPosition" AT %ID2904 : DWord;   // CARRIER POSITION
   "Carrier_51_CarrierNumber" AT %IW2908 : Word;   // CARRIER NUMBER
   "Carrier_51_G120DControlWord" AT %IW2910 : Word;   // G120D_STW1_CONTROL
   "Carrier_51_G120DControlWord.0" AT %I2910.0 : Bool;   // Bit_00_ON
   "Carrier_51_G120DControlWord.1" AT %I2910.1 : Bool;   // Bit_01_AUS2_INH
   "Carrier_51_G120DControlWord.2" AT %I2910.2 : Bool;   // Bit_02_AUS3_STOP
   "Carrier_51_G120DControlWord.3" AT %I2910.3 : Bool;   // Bit_03_EN
   "Carrier_51_G120DControlWord.4" AT %I2910.4 : Bool;   // Bit_04_EN_RAMP
   "Carrier_51_G120DControlWord.5" AT %I2910.5 : Bool;   // Bit_05_START_RAMP
   "Carrier_51_G120DControlWord.6" AT %I2910.6 : Bool;   // Bit_06_SETPOINT
   "Carrier_51_G120DControlWord.7" AT %I2910.7 : Bool;   // Bit_07_RESET
   "Carrier_51_G120DControlWord.8" AT %I2911.0 : Bool;   // Bit_08_JOG_R
   "Carrier_51_G120DControlWord.9" AT %I2911.1 : Bool;   // Bit_09_JOG_L
   "Carrier_51_G120DControlWord.10" AT %I2911.2 : Bool;   // Bit_10_CONTR_PLC
   "Carrier_51_G120DControlWord.11" AT %I2911.3 : Bool;   // Bit_11_REVERSE
   "Carrier_51_G120DControlWord.12" AT %I2911.4 : Bool;   // Bit_12_BRAKE_RELEASE
   "Carrier_51_G120DControlWord.13" AT %I2911.5 : Bool;   // Bit_13_DDS
   "Carrier_51_G120DControlWord.14" AT %I2911.6 : Bool;   // Bit_14_DO0
   "Carrier_51_G120DControlWord.15" AT %I2911.7 : Bool;   // Bit_15_DO1
   "Carrier_51_G120DStatusWord" AT %IW2912 : Word;   // G120D_ZSW1_STATUS